(* CODESYS project Revisora_V2.0.1h.project (continued)
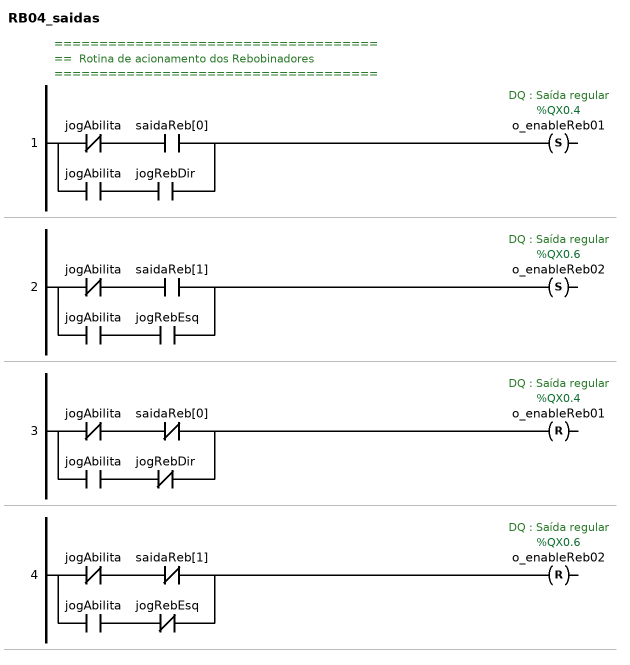
// NETWORK 1
// ====================================
// ==  Rotina de acionamento dos Rebobinadores
// ====================================
//   o_enableReb01: DQ : Saída regular | AT %QX0.4
o_enableReb01 S= NOT jogAbilita AND saidaReb[0] OR jogAbilita AND jogRebDir;

// NETWORK 2
//   o_enableReb02: DQ : Saída regular | AT %QX0.6
o_enableReb02 S= NOT jogAbilita AND saidaReb[1] OR jogAbilita AND jogRebEsq;

// NETWORK 3
//   o_enableReb01: DQ : Saída regular | AT %QX0.4
o_enableReb01 R= NOT jogAbilita AND NOT saidaReb[0] OR jogAbilita AND NOT jogRebDir;

// NETWORK 4
//   o_enableReb02: DQ : Saída regular | AT %QX0.6
o_enableReb02 R= NOT jogAbilita AND NOT saidaReb[1] OR jogAbilita AND NOT jogRebEsq;

END_PROGRAM

// MyController/Application/02_Rebobinadores/RB05_sentido
PROGRAM RB05_sentido
VAR
auxParseAnalog				:ARRAY [1..2] OF REAL;
END_VAR

// Calcula quando o valor for menor que 0
auxParseAnalog[1]:= (parseAnalog[0] * 100) / 1;
auxParseAnalog[2]:= (parseAnalog[1] * 100) / 1;



//IF parseAnalog[0] < 0 THEN
	//valorPorcRebobinador[1]:= auxParseAnalog[1];
//ELSE
	//valorPorcRebobinador[1]:= porcRebobinador[1];	
//END_IF

IF parseAnalog[1] < 0 THEN
	valorPorcRebobinador[2]:= auxParseAnalog[2];
ELSE
	valorPorcRebobinador[2]:= porcRebobinador[2];	
END_IF

// Sentido dos rebobinadores
IF	enbReb.IP THEN
	IF i_sentido THEN
		ladoDir:= FALSE;
		ladoEsq:= TRUE;
		visLadoEsq:= TRUE;
		visLadoDir:= FALSE;
		displayState:= 0;
	ELSE
		ladoEsq:= FALSE;
		ladoDir:= TRUE;
		visLadoEsq:= FALSE;
		visLadoDir:= TRUE;
		displayState:= 1;
	END_IF
END_IF

// Editar valores

	IF ladoEsq THEN
		oa_saidaTorque_2:= REAL_TO_INT((auxParseAnalog[1])*-1); 
		oa_saidaTorque_1:= REAL_TO_INT((auxParseAnalog[2]));
		delayTorq[0] := T#500MS;
		delayTorq[1] := T#0MS;
		
	END_IF
	
	IF ladoDir THEN
		oa_saidaTorque_2:= REAL_TO_INT(auxParseAnalog[2])*-1;
		oa_saidaTorque_1:= REAL_TO_INT(auxParseAnalog[1]);
		delayTorq[0] := T#0MS;
		delayTorq[1] := T#500MS;
	END_IF
	
	//IF NOT ciclo.IP THEN
	//	ladoEsq:= FALSE;
	//	ladoDir:= FALSE;
//	END_IF
	
	// Parada
	IF torqueParada THEN
		IF ladoEsq THEN
			oa_saidaTorque_2:= 1311;
			oa_saidaTorque_1:= 5000;
		ELSE
			oa_saidaTorque_2:= -5000;
			oa_saidaTorque_1:= -1311;
		END_IF
	END_IF
// Calcula quando o valor for menor que 0
//auxParseAnalog[1]:= (parseAnalog[0] * 328) / 3;
//auxParseAnalog[2]:= (parseAnalog[1] * 328) / 3;

END_PROGRAM

// MyController/Application/03_Nip/NP01_geral
PROGRAM NP01_geral
VAR
	TD_power				: TOF;
END_VAR
VAR // added by the converter: edge detectors and wires of the graphical bodies
    _ft1 : F_TRIG;
END_VAR

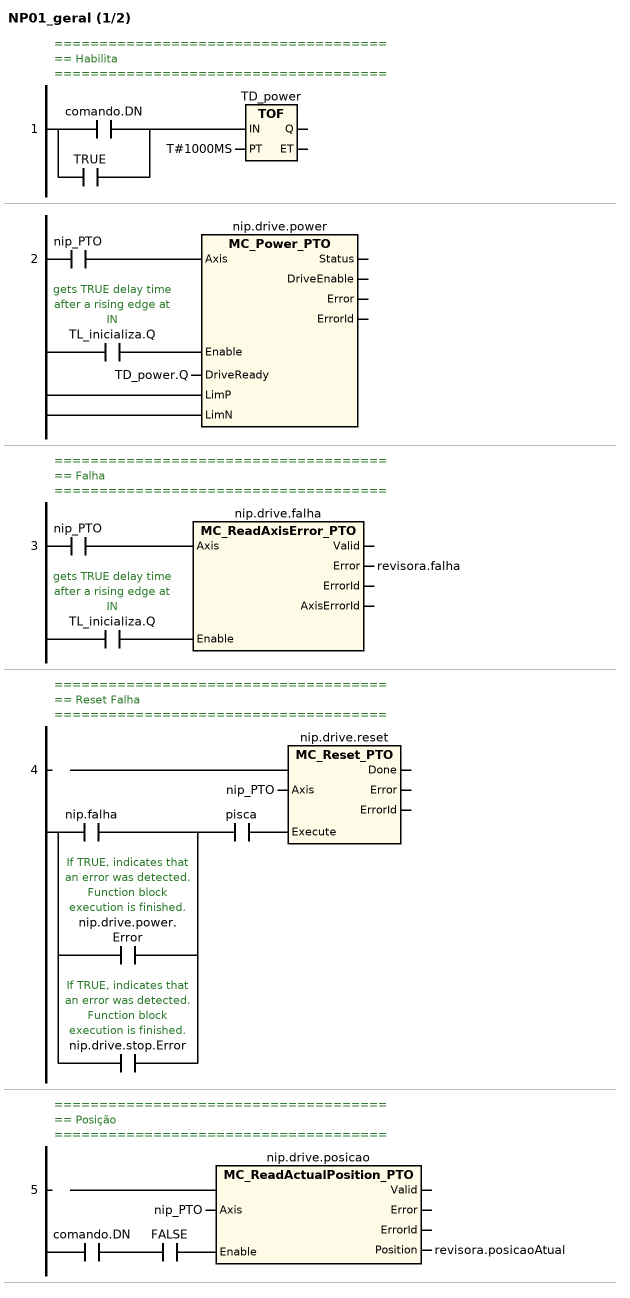
// NETWORK 1
// =====================================
// == Habilita
// =====================================
TD_power(IN := comando.DN OR TRUE, PT := T#1000MS); // TOF

// NETWORK 2
//   TL_inicializa.Q: gets TRUE delay time after a rising edge at IN
//   TD_power.Q: gets FALSE, when PT milliseconds elapsed, since falling edge at IN
nip.drive.power(
    Axis := nip_PTO,
    Enable := TL_inicializa.Q,
    DriveReady := TD_power.Q,
    LimP := TRUE,
    LimN := TRUE); // MC_Power_PTO

// NETWORK 3
// =====================================
// == Falha
// =====================================
//   TL_inicializa.Q: gets TRUE delay time after a rising edge at IN
nip.drive.falha(Axis := nip_PTO, Enable := TL_inicializa.Q, Error => revisora.falha); // MC_ReadAxisError_PTO

// NETWORK 4
// =====================================
// == Reset Falha
// =====================================
//   nip.drive.power.Error: If TRUE, indicates that an error was detected. Function block execution is finished.
//   nip.drive.stop.Error: If TRUE, indicates that an error was detected. Function block execution is finished.
nip.drive.reset(Axis := nip_PTO, Execute := (nip.falha OR nip.drive.power.Error OR nip.drive.stop.Error) AND pisca); // MC_Reset_PTO

// NETWORK 5
// =====================================
// == Posição
// =====================================
nip.drive.posicao(Axis := nip_PTO, Enable := comando.DN AND FALSE, Position => revisora.posicaoAtual); // MC_ReadActualPosition_PTO

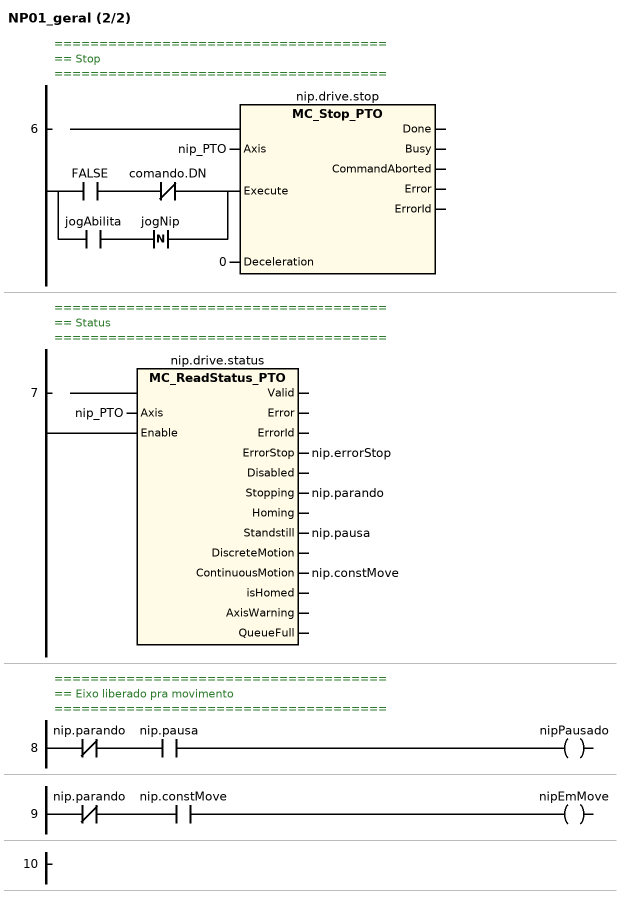
// NETWORK 6
// =====================================
// == Stop
// =====================================
_ft1(CLK := jogNip);
nip.drive.stop(
    Axis := nip_PTO,
    Execute := FALSE AND NOT comando.DN OR jogAbilita AND _ft1.Q,
    Deceleration := 0); // MC_Stop_PTO

// NETWORK 7
// =====================================
// == Status
// =====================================
nip.drive.status(
    Axis := nip_PTO,
    Enable := TRUE,
    ErrorStop => nip.errorStop,
    Stopping => nip.parando,
    Standstill => nip.pausa,
    ContinuousMotion => nip.constMove); // MC_ReadStatus_PTO

// NETWORK 8
// =====================================
// == Eixo liberado pra movimento
// =====================================
nipPausado := NOT nip.parando AND nip.pausa;

// NETWORK 9
nipEmMove := NOT nip.parando AND nip.constMove;

// NETWORK 10

END_PROGRAM

// MyController/Application/03_Nip/NP02_enableNip
PROGRAM NP02_enableNip
VAR
END_VAR

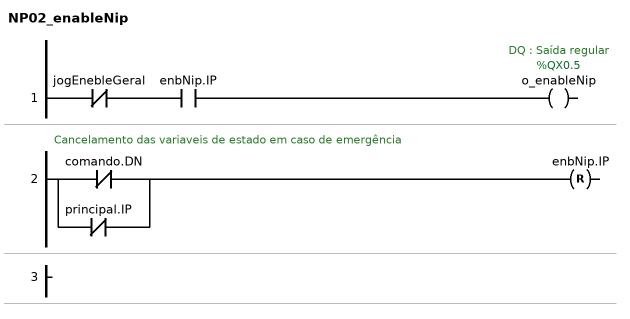
// NETWORK 1
//   o_enableNip: DQ : Saída regular | AT %QX0.5
o_enableNip := NOT jogEnebleGeral AND enbNip.IP;

// NETWORK 2
// Cancelamento das variaveis de estado em caso de emergência
enbNip.IP R= NOT comando.DN OR NOT principal.IP;

// NETWORK 3

END_PROGRAM

// MyController/Application/03_Nip/NP03_auto
PROGRAM NP03_auto
VAR
	TF_enable						: TON;
	MC_MoveVelocity_PTO_0			: MC_MoveVelocity_PTO;
	atrasoAposDesligar				: ARRAY [1..2] OF TON;
	testeTempo: TP;
END_VAR
VAR // added by the converter: edge detectors and wires of the graphical bodies
    _ft1, _ft2, _ft3 : F_TRIG;
    _rt1 : R_TRIG;
    _w1, _w2 : BOOL;
END_VAR

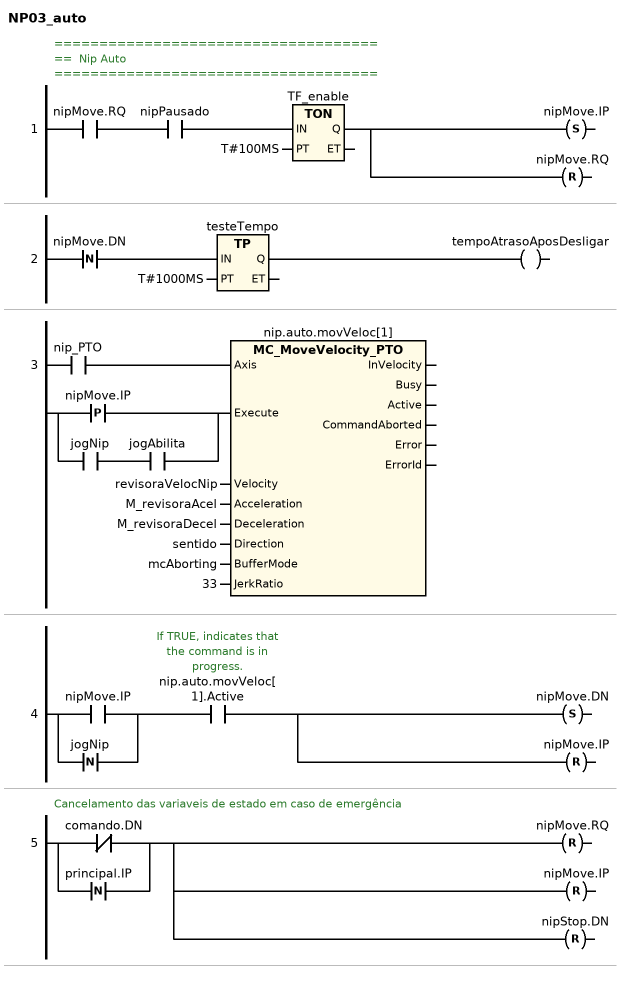
// NETWORK 1
// ====================================
// ==  Nip Auto
// ====================================
TF_enable(IN := nipMove.RQ AND nipPausado, PT := T#100MS); // TON
nipMove.IP S= TF_enable.Q;
nipMove.RQ R= TF_enable.Q;

// NETWORK 2
_ft1(CLK := nipMove.DN);
testeTempo(IN := _ft1.Q, PT := T#1000MS); // TP
tempoAtrasoAposDesligar := testeTempo.Q;

// NETWORK 3
_rt1(CLK := nipMove.IP);
nip.auto.movVeloc[1](
    Axis := nip_PTO,
    Execute := _rt1.Q OR jogNip AND jogAbilita,
    Velocity := revisoraVelocNip,
    Acceleration := M_revisoraAcel,
    Deceleration := M_revisoraDecel,
    Direction := sentido,
    BufferMode := mcAborting,
    JerkRatio := 33); // MC_MoveVelocity_PTO

// NETWORK 4
//   nip.auto.movVeloc[1].Active: If TRUE, indicates that the command is in progress.
_ft2(CLK := jogNip);
_w1 := (nipMove.IP OR _ft2.Q) AND nip.auto.movVeloc[1].Active;
nipMove.DN S= _w1;
nipMove.IP R= _w1;

// NETWORK 5
// Cancelamento das variaveis de estado em caso de emergência
_ft3(CLK := principal.IP);
_w2 := NOT comando.DN OR _ft3.Q;
nipMove.RQ R= _w2;
nipMove.IP R= _w2;
nipStop.DN R= _w2;

END_PROGRAM

// MyController/Application/03_Nip/NP04_parada
PROGRAM NP04_parada
VAR
	testeFW			: BOOL;
	job: BOOL;
	atradoZeraPosicao: TON;
END_VAR
VAR // added by the converter: edge detectors and wires of the graphical bodies
    _w1, _w2, _w3 : BOOL;
    _rt1 : R_TRIG;
    _ft1 : F_TRIG;
END_VAR

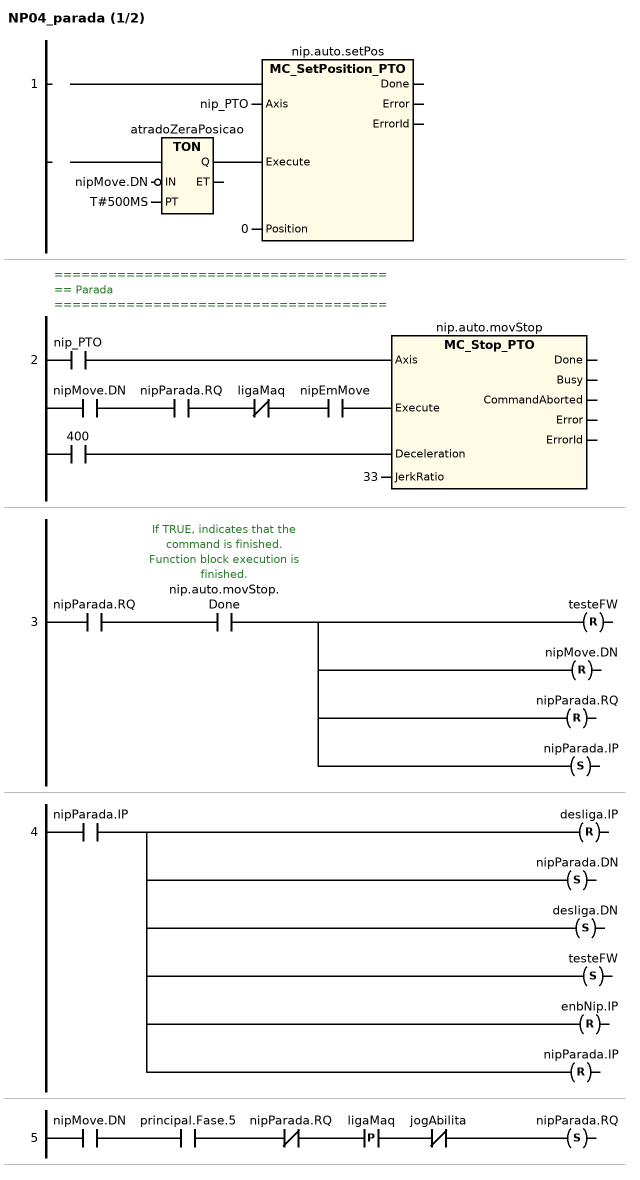
// NETWORK 1
atradoZeraPosicao(IN := NOT nipMove.DN, PT := T#500MS); // TON
nip.auto.setPos(Axis := nip_PTO, Execute := atradoZeraPosicao.Q, Position := 0); // MC_SetPosition_PTO

// NETWORK 2
// =====================================
// == Parada
// =====================================
nip.auto.movStop(
    Axis := nip_PTO,
    Execute := nipMove.DN AND nipParada.RQ AND NOT ligaMaq AND nipEmMove,
    Deceleration := 400,
    JerkRatio := 33); // MC_Stop_PTO

// NETWORK 3
//   nip.auto.movStop.Done: If TRUE, indicates that the command is finished. Function block execution is finished.
_w1 := nipParada.RQ AND nip.auto.movStop.Done;
testeFW R= _w1;
nipMove.DN R= _w1;
nipParada.RQ R= _w1;
nipParada.IP S= _w1;

// NETWORK 4
_w2 := nipParada.IP;
desliga.IP R= _w2;
nipParada.DN S= _w2;
desliga.DN S= _w2;
testeFW S= _w2;
enbNip.IP R= _w2;
nipParada.IP R= _w2;

// NETWORK 5
_rt1(CLK := ligaMaq);
nipParada.RQ S= nipMove.DN AND principal.Fase.5 AND NOT nipParada.RQ AND _rt1.Q AND NOT jogAbilita;

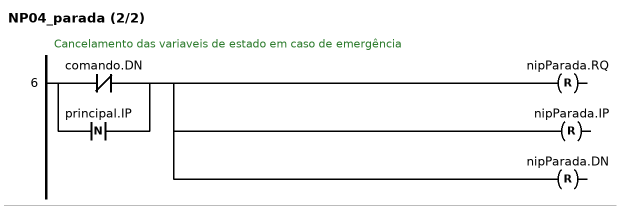
// NETWORK 6
// Cancelamento das variaveis de estado em caso de emergência
_ft1(CLK := principal.IP);
_w3 := NOT comando.DN OR _ft1.Q;
nipParada.RQ R= _w3;
nipParada.IP R= _w3;
nipParada.DN R= _w3;

END_PROGRAM

// MyController/Application/03_Nip/NP06_jog
PROGRAM NP06_jog
VAR
	auxJogPos								: BOOL;
	auxJopNeg								: BOOL;
END_VAR
VAR // added by the converter: edge detectors and wires of the graphical bodies
    _ft1, _ft2 : F_TRIG;
END_VAR

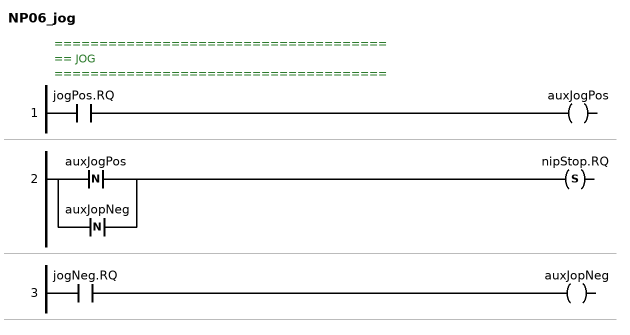
// NETWORK 1
// =====================================
// == JOG
// =====================================
auxJogPos := jogPos.RQ;

// NETWORK 2
_ft1(CLK := auxJogPos);
_ft2(CLK := auxJopNeg);
nipStop.RQ S= _ft1.Q OR _ft2.Q;

// NETWORK 3
auxJopNeg := jogNeg.RQ;

END_PROGRAM

// MyController/Application/03_Nip/NP07_veloc
PROGRAM NP07_veloc
VAR

	timerVeloc 		: TON;

END_VAR

// Partida Lenta
IF sentido = -1 THEN
	M_revisoraVeloc:=bobinaAtual.velocReb;
END_IF
IF sentido = 1 THEN
	M_revisoraVeloc:=bobinaAtual.velocDesb;
END_IF
//IF nipMove.RQ THEN
//	IF bobinaAtual.velocDesb > 800 OR bobinaAtual.velocReb > 800 THEN	
	//	M_revisoraVeloc:= 600;
	//	partidaLenta:= TRUE;
//	END_IF
//END_IF

//timerVeloc(IN:= partidaLenta, PT:= T#7S);

//IF 	timerVeloc.Q THEN
	//nipMove.IP:= FALSE;
	//partidaLenta:= FALSE;
	//IF i_sentido THEN
	//	M_revisoraVeloc:= bobinaAtual.velocDesb;
	//	nipMove.IP:= TRUE;
//	ELSE
//		M_revisoraVeloc:= bobinaAtual.velocReb;
//		nipMove.IP:= TRUE;
//	END_IF
//END_IF

//IF NOT comando.DN OR principal.IP OR ligaMaq THEN
//	partidaLenta:= FALSE;
//END_IF

END_PROGRAM

// MyController/Application/03_Nip/NP09_sentido
PROGRAM NP09_sentido
VAR
END_VAR

// Mudança de sentido
IF i_sentido AND NOT ciclo.IP THEN
	sentido:= 1;
	M_pulsosParar:= 20;
ELSIF NOT i_sentido AND NOT ciclo.IP THEN
	sentido:= -1;
	M_pulsosParar:= -20;
END_IF

END_PROGRAM

// MyController/Application/03_Nip/NP20_JogTest
PROGRAM NP20_JogTest
VAR
	auxVeloc			:DINT;
	auxReb01			: INT;
	auxReb02			: INT;
END_VAR

IF jogVelocNip >3000 THEN
	jogVelocNip:= 3000;
	
END_IF

IF jogAbilita = TRUE THEN
	revisoraVelocNip:=jogVelocNip;
ELSE
	revisoraVelocNip:=M_revisoraVeloc;
END_IF

END_PROGRAM

// MyController/Application/05_IHM/I01_geral
PROGRAM I01_geral
VAR
	auxBit				: BOOL;
END_VAR
VAR // added by the converter: edge detectors and wires of the graphical bodies
    _rt1 : R_TRIG;
END_VAR

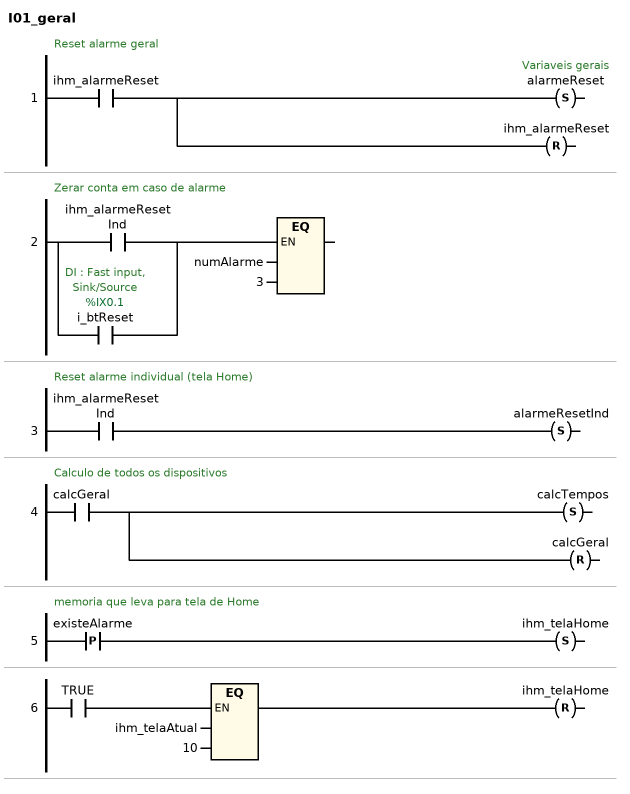
// NETWORK 1
// Reset alarme geral
//   alarmeReset: Variaveis gerais
alarmeReset S= ihm_alarmeReset;
ihm_alarmeReset R= ihm_alarmeReset;

// NETWORK 2
// Zerar conta em caso de alarme
//   i_btReset: DI : Fast input, Sink/Source | AT %IX0.1
(* (ihm_alarmeResetInd OR i_btReset) AND numAlarme = 3; result not used *)

// NETWORK 3
// Reset alarme individual (tela Home)
alarmeResetInd S= ihm_alarmeResetInd;

// NETWORK 4
// Calculo de todos os dispositivos
calcTempos S= calcGeral;
calcGeral R= calcGeral;

// NETWORK 5
// memoria que leva para tela de Home
_rt1(CLK := existeAlarme);
ihm_telaHome S= _rt1.Q;

// NETWORK 6
ihm_telaHome R= ihm_telaAtual = 10;

END_PROGRAM

// MyController/Application/05_IHM/I02_alarmes
PROGRAM I02_alarmes
VAR
	auxExisteAlarme					: BOOL;
	delayAlarme						: TON;
	memAlarme						: ARRAY[0..99] OF BOOL;
	p0								: SINT;
END_VAR


CASE alarmes.Fase OF
(*====================================
  ==  Fase 0 - alarmes 1 a 50 (0 não existe)
  ====================================*)
0:
	auxExisteAlarme:= FALSE;
	FOR p0:= 1 TO 50 DO
		IF alarme[p0] THEN
			memAlarme[p0]:= TRUE;
			auxExisteAlarme:= TRUE;
			
			IF numAlarme = 0 THEN
				numAlarme:= p0;				// pega o numero do primeiro alarme que ocorre
			END_IF
		END_IF
		
		IF numAlarme = p0 THEN
			IF alarme[p0] = 0 THEN			// verifica se o alarme que ocorreu continua ativo
				numAlarme:= 0;
			END_IF
		END_IF
	END_FOR
	alarmes.Fase:= 10;

	
(*====================================
  ==  Fase 10 - passa alarmes para ihm	
  ====================================*)
10:
	FOR p0:= 1 TO 50 DO
		ihm_alarme[p0]:= memAlarme[p0];
		memAlarme[p0]:= FALSE;
	END_FOR
	alarmes.Fase:= 11;
	
	
(*====================================
  ==  Fase 11 - verifica cancela alarmes pela IHM
  ====================================*)	
11:
	existeAlarme:= auxExisteAlarme;
	IF alarmeReset THEN
		alarmes.Fase:= 12;
	ELSE
		IF alarmeResetInd OR (i_btReset AND comando.DN) THEN
			alarme[numAlarme]:= FALSE;
			alarmeResetInd:= FALSE;
		END_IF
		alarmes.Fase:= 0;
	END_IF

	
(*====================================
  ==  Fase 12 - cancela alarmes	
  ====================================*)
12:
	alarmeReset:= FALSE;
	FOR p0:= 1 TO 50 DO
		alarme[p0]:= 0;
	END_FOR
	alarmes.Fase:= 13;
	

(*====================================
  ==  Fase 13 - espera 100ms para atualização dos bits de alarmes pelo controle
  ====================================*)	
13:
	IF delayAlarme.Q THEN
		alarmes.Fase:= 0;
	END_IF
	delayAlarme(IN:= alarmes.Fase= 13, PT:= T#100MS);

END_CASE

END_PROGRAM

// MyController/Application/05_IHM/I03_mensagens
PROGRAM I03_mensagens
VAR
	delayMensag						: TON;
	mensagens						: _exec_bits;
	p1								: DINT;
END_VAR


IF NOT mensagens.RQ THEN
	FOR p1:= 1 TO 50 DO
		IF mensagem[p1] = TRUE THEN
			mensagem[p1]:= 0;
			ihm_mensagem:= p1;
			mensagens.RQ:= TRUE;
		END_IF
	END_FOR
END_IF


// Tempo de cada mensagem na tela
delayMensag(IN := ihm_bannerMensagem, PT:= T#2500MS);
IF delayMensag.Q THEN
	mensagens.RQ:= FALSE;
	ihm_mensagem:= 0;
END_IF


ihm_bannerMensagem:= mensagens.RQ AND NOT ihm_bannerConfirma;

END_PROGRAM

// MyController/Application/05_IHM/I06_textoConfirma
PROGRAM I06_textoConfirma
VAR
END_VAR
VAR // added by the converter: edge detectors and wires of the graphical bodies
    _w1 : BOOL;
END_VAR

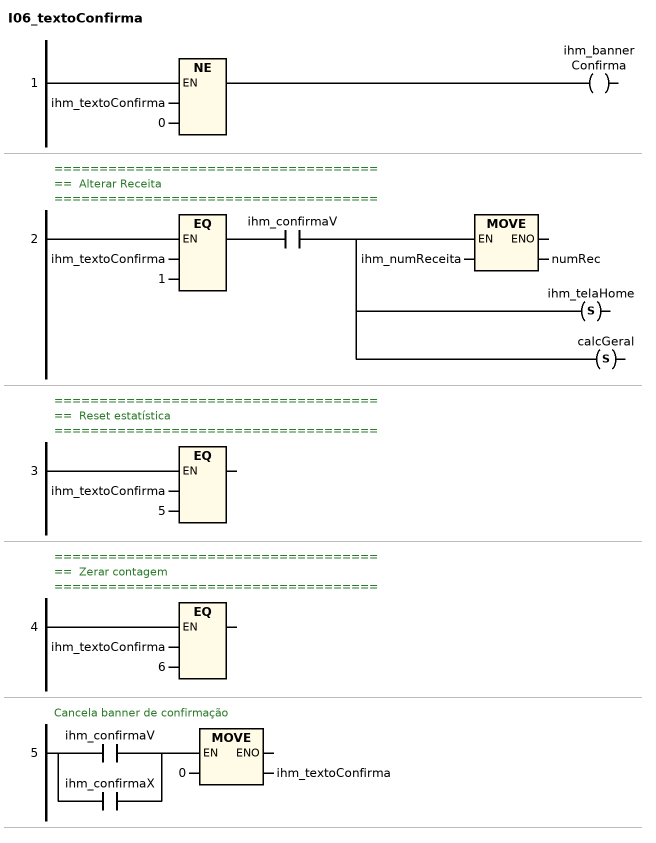
// NETWORK 1
ihm_bannerConfirma := ihm_textoConfirma <> 0;

// NETWORK 2
// ====================================
// ==  Alterar Receita
// ====================================
_w1 := ihm_textoConfirma = 1 AND ihm_confirmaV;
IF _w1 THEN numRec := ihm_numReceita; END_IF
ihm_telaHome S= _w1;
calcGeral S= _w1;

// NETWORK 3
// ====================================
// ==  Reset estatística
// ====================================
(* ihm_textoConfirma = 5; result not used *)

// NETWORK 4
// ====================================
// ==  Zerar contagem
// ====================================
(* ihm_textoConfirma = 6; result not used *)

// NETWORK 5
// Cancela banner de confirmação
IF ihm_confirmaV OR ihm_confirmaX THEN ihm_textoConfirma := 0; END_IF

END_PROGRAM

// MyController/Application/19_Ultrassonico/U10_auto
PROGRAM U10_auto
VAR

END_VAR
VAR // added by the converter: edge detectors and wires of the graphical bodies
    _rt1, _rt2, _rt3, _rt4 : R_TRIG;
END_VAR

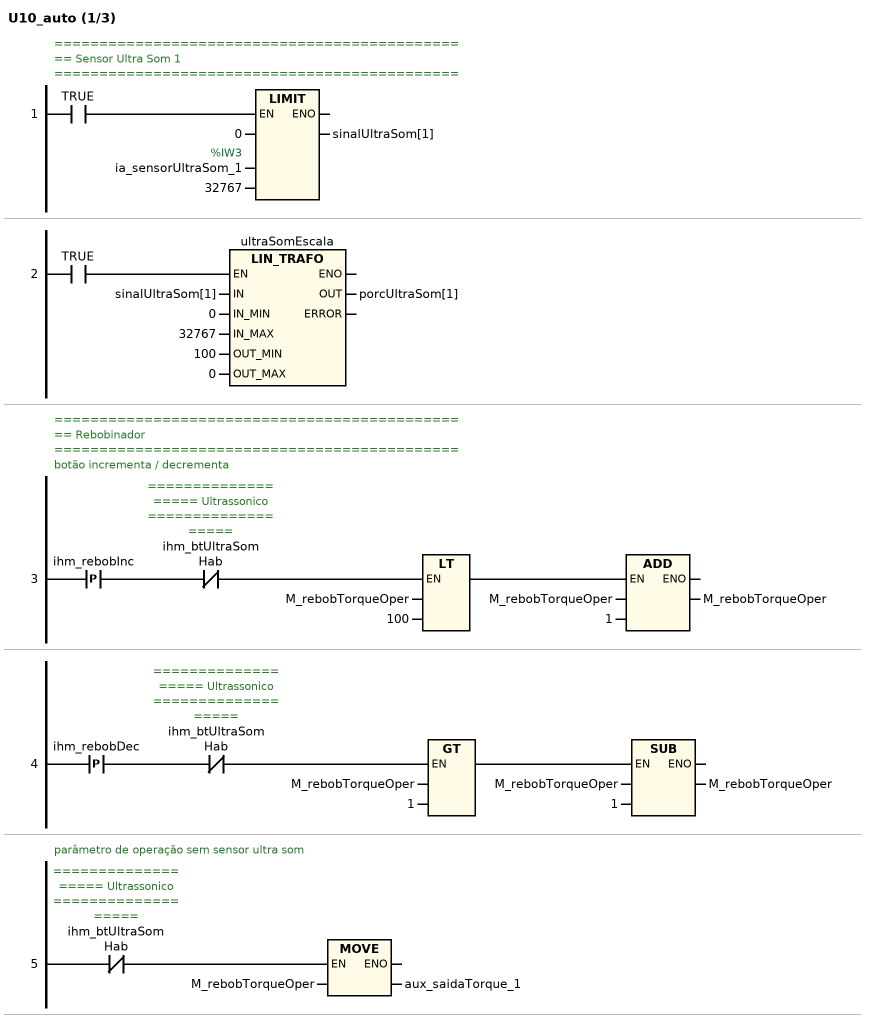
// NETWORK 1
// =============================================
// == Sensor Ultra Som 1
// =============================================
//   ia_sensorUltraSom_1: Ultra : | AT %IW3
sinalUltraSom[1] := LIMIT(0, ia_sensorUltraSom_1, 32767);

// NETWORK 2
ultraSomEscala(
    IN := sinalUltraSom[1],
    IN_MIN := 0,
    IN_MAX := 32767,
    OUT_MIN := 100,
    OUT_MAX := 0,
    OUT => porcUltraSom[1]); // LIN_TRAFO

// NETWORK 3
// =============================================
// == Rebobinador
// =============================================
// botão incrementa / decrementa
//   ihm_btUltraSomHab: =================== Ultrassonico ===================
_rt1(CLK := ihm_rebobInc);
IF _rt1.Q AND NOT ihm_btUltraSomHab AND M_rebobTorqueOper < 100 THEN
    M_rebobTorqueOper := M_rebobTorqueOper + 1;
END_IF

// NETWORK 4
//   ihm_btUltraSomHab: =================== Ultrassonico ===================
_rt2(CLK := ihm_rebobDec);
IF _rt2.Q AND NOT ihm_btUltraSomHab AND M_rebobTorqueOper > 1 THEN
    M_rebobTorqueOper := M_rebobTorqueOper - 1;
END_IF

// NETWORK 5
// parâmetro de operação sem sensor ultra som
//   ihm_btUltraSomHab: =================== Ultrassonico ===================
//   aux_saidaTorque_1: =================== Ultrassonico =================== ia_sensorUltraSom_1 :INT; ia_sensorUltraSom_2 :INT;
IF NOT ihm_btUltraSomHab THEN aux_saidaTorque_1 := M_rebobTorqueOper; END_IF

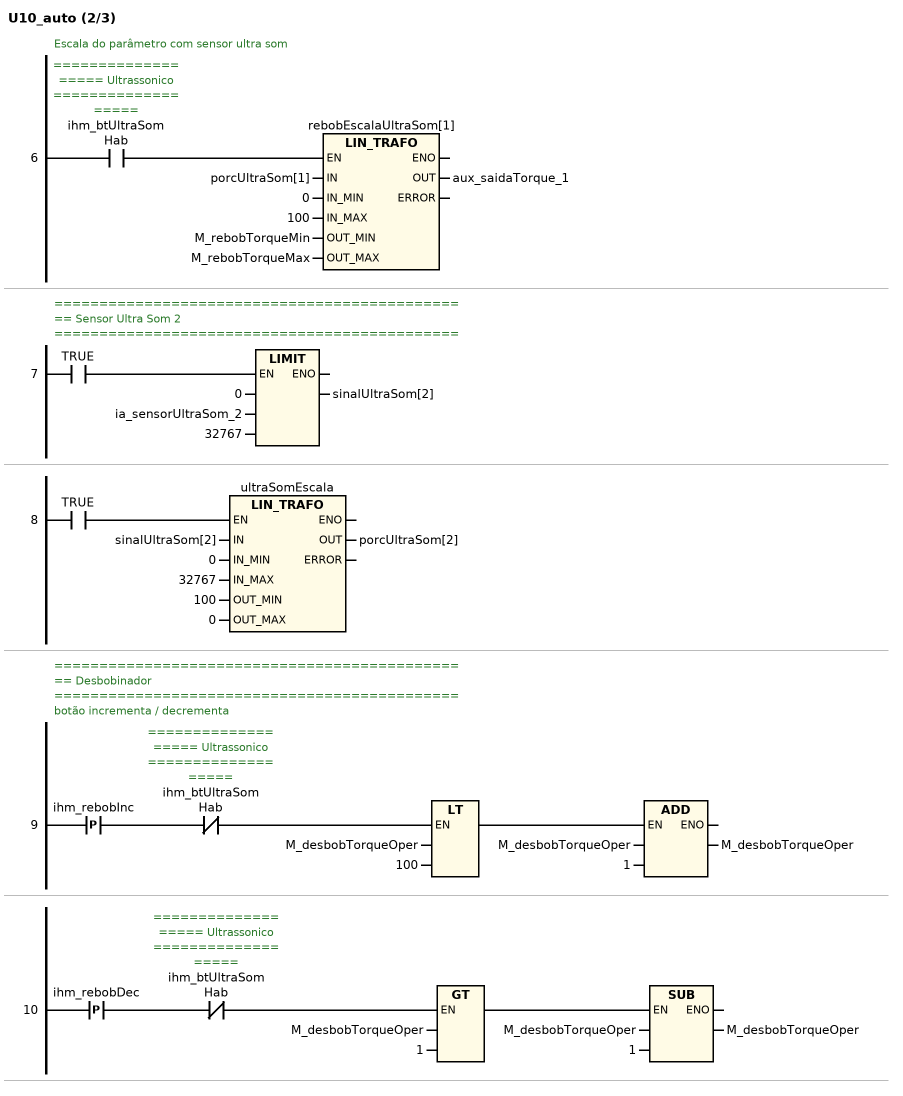
// NETWORK 6
// Escala do parâmetro com sensor ultra som
//   ihm_btUltraSomHab: =================== Ultrassonico ===================
//   aux_saidaTorque_1: =================== Ultrassonico =================== ia_sensorUltraSom_1 :INT; ia_sensorUltraSom_2 :INT;
IF ihm_btUltraSomHab THEN
    rebobEscalaUltraSom[1](
        IN := porcUltraSom[1],
        IN_MIN := 0,
        IN_MAX := 100,
        OUT_MIN := M_rebobTorqueMin,
        OUT_MAX := M_rebobTorqueMax,
        OUT => aux_saidaTorque_1); // LIN_TRAFO
END_IF

// NETWORK 7
// =============================================
// == Sensor Ultra Som 2
// =============================================
sinalUltraSom[2] := LIMIT(0, ia_sensorUltraSom_2, 32767);

// NETWORK 8
ultraSomEscala(
    IN := sinalUltraSom[2],
    IN_MIN := 0,
    IN_MAX := 32767,
    OUT_MIN := 100,
    OUT_MAX := 0,
    OUT => porcUltraSom[2]); // LIN_TRAFO

// NETWORK 9
// =============================================
// == Desbobinador
// =============================================
// botão incrementa / decrementa
//   ihm_btUltraSomHab: =================== Ultrassonico ===================
_rt3(CLK := ihm_rebobInc);
IF _rt3.Q AND NOT ihm_btUltraSomHab AND M_desbobTorqueOper < 100 THEN
    M_desbobTorqueOper := M_desbobTorqueOper + 1;
END_IF

// NETWORK 10
//   ihm_btUltraSomHab: =================== Ultrassonico ===================
_rt4(CLK := ihm_rebobDec);
IF _rt4.Q AND NOT ihm_btUltraSomHab AND M_desbobTorqueOper > 1 THEN
    M_desbobTorqueOper := M_desbobTorqueOper - 1;
END_IF

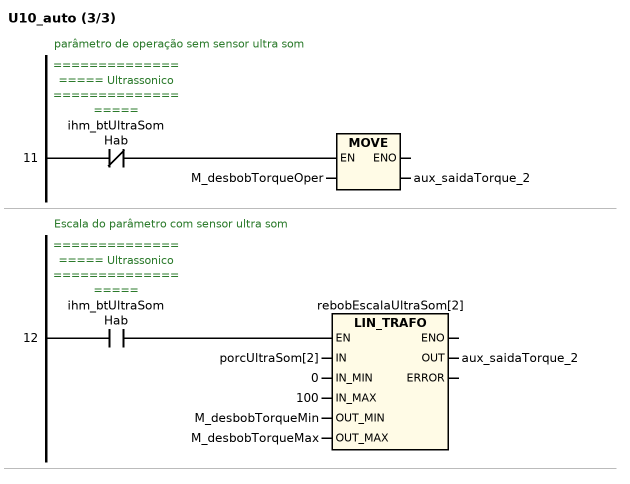
// NETWORK 11
// parâmetro de operação sem sensor ultra som
//   ihm_btUltraSomHab: =================== Ultrassonico ===================
IF NOT ihm_btUltraSomHab THEN aux_saidaTorque_2 := M_desbobTorqueOper; END_IF

// NETWORK 12
// Escala do parâmetro com sensor ultra som
//   ihm_btUltraSomHab: =================== Ultrassonico ===================
IF ihm_btUltraSomHab THEN
    rebobEscalaUltraSom[2](
        IN := porcUltraSom[2],
        IN_MIN := 0,
        IN_MAX := 100,
        OUT_MIN := M_desbobTorqueMin,
        OUT_MAX := M_desbobTorqueMax,
        OUT => aux_saidaTorque_2); // LIN_TRAFO
END_IF

END_PROGRAM

// MyController/Application/19_Ultrassonico/U99_calculo
PROGRAM U99_calculo
VAR
END_VAR

// Envia valores

oa_saidaTorque_1:= REAL_TO_INT(aux_saidaTorque_1);
oa_saidaTorque_2:= REAL_TO_INT(aux_saidaTorque_2);

END_PROGRAM

// MyController/Application/10_Relogio/AjustaDataHora
PROGRAM AjustaDataHora
VAR
	writeDateTime			: SetDateAndTime;
	readDateTime			: GetDateAndTime;
	bitScan					: BOOL;
	comOk					: BOOL;
	T_com					: TON;
END_VAR
VAR // added by the converter: edge detectors and wires of the graphical bodies
    _rt1 : R_TRIG;
END_VAR

